
                   IF #AUX_tFM152RecvAck.bACK = #CONST_BFM152_ACK THEN
                       #TMP_xFm152ValidReply := TRUE;
                   END_IF;
               END_IF;

           #CONST_DFM152_TEL_WRITERAMPJOG:        

               IF #AUX_dActualElBuffer = #CONST_DFM152_ACK_NACKSIZE THEN

                   #TMP_dBufferPos := 0;
                   #TMP_iRetVal := Deserialize(SRC_ARRAY:=#AUX_rgbReceiveBuffer, DEST_VARIABLE=>#AUX_tFM152RecvAck, POS:=#TMP_dBufferPos);

                   IF #AUX_tFM152RecvAck.bACK = #CONST_BFM152_ACK THEN
                       #TMP_xFm152ValidReply := TRUE;
                   END_IF;
               END_IF;

           #CONST_DFM152_TEL_WRITERAMP:        

               IF #AUX_dActualElBuffer = #CONST_DFM152_ACK_NACKSIZE THEN

                   #TMP_dBufferPos := 0;
                   #TMP_iRetVal := Deserialize(SRC_ARRAY:=#AUX_rgbReceiveBuffer, DEST_VARIABLE=>#AUX_tFM152RecvAck, POS:=#TMP_dBufferPos);

                   IF #AUX_tFM152RecvAck.bACK = #CONST_BFM152_ACK THEN
                       #TMP_xFm152ValidReply := TRUE;
                   END_IF;
               END_IF;

           #CONST_DFM152_TEL_REQACTDATA: 

               IF #AUX_dActualElBuffer = #CONST_DFM152_ACK_NACKSIZE THEN

                   #TMP_dBufferPos := 0;
                   #TMP_iRetVal := Deserialize(SRC_ARRAY:=#AUX_rgbReceiveBuffer, DEST_VARIABLE=>#AUX_tFM152RecvAck, POS:=#TMP_dBufferPos);

                   IF #AUX_tFM152RecvAck.bACK = #CONST_BFM152_ACK THEN
                       #TMP_xFm152ValidReply := TRUE;
                   END_IF;
               END_IF;

       END_CASE;

       IF #TMP_xFm152ValidReply = TRUE THEN
           #AUX_dActualElBuffer := 0;
       END_IF;

   ELSE
       #AUX_dActualElBuffer := 0;
   END_IF;
END_REGION

REGION Network 39: End waiting data reply
   RUNG wire#powerrail
      Contact( #tPhases.xWaitingFm152Reply )
      wire#w1
      Contact( #TMP_xFm152ValidReply )
      wire#w2
      R_Coil( #tPhases.xWaitingFm152Reply )
   END_RUNG
   RUNG wire#w1
      Contact( #tmON_TimeoutRecvData.Q )
   END_RUNG wire#w2
   RUNG wire#w2
      Coil( #tPhases.xEndWaitingFm152Reply )
   END_RUNG
   // the same network as SCL:
   #_w1 := #tPhases.xWaitingFm152Reply AND (#TMP_xFm152ValidReply OR #tmON_TimeoutRecvData.Q);
   IF #_w1 THEN #tPhases.xWaitingFm152Reply := FALSE; END_IF;
   #tPhases.xEndWaitingFm152Reply := #_w1;
END_REGION

REGION Network 40 (SCL): Phase in progress
   GATHER(IN:=#tPhases,
          OUT=>#TMP_dwValue);

   IF #TMP_dwValue <> 0 THEN
       #ST_xFm152PhaseProgr := TRUE;
   ELSE
       #ST_xFm152PhaseProgr := FALSE;
   END_IF;
END_REGION
END_FUNCTION_BLOCK

FUNCTION_BLOCK "FB_DigitizerManager_V1.00"   // FB4, LAD
{ S7_Optimized_Access := 'TRUE' }
VERSION : 0.1
   VAR_INPUT
      IN_xCycleON : Bool;   // Cycle ON
      IN_xCycleONDel : Bool;   // Delayed cycle ON signal
      IN_xGeneralReset : Bool;   // General reset
      IN_xResetAlarms : Bool;   // Reset alarms
      IN_xFaultsEnabled : Bool;   // Faults enabled
   END_VAR
   VAR_OUTPUT
      OUTPUTS : Struct   // OUTPUTS
         xEnableJog : Bool;   // OUTPUT.Enable jog
         xSelectEncoder1 : Bool;   // OUTPUT.Select encoder #1
      END_STRUCT;
   END_VAR
   VAR_IN_OUT
      INO_tDigitizer1 : "FB_Digitizer_V1.00";   // Digitizer #1
      INO_tDigitizer2 : "FB_Digitizer_V1.00";   // Digitizer #2
      INO_tEnc : "UDT_Encoder";   // Encoder
   END_VAR
   VAR RETAIN
      tHMR : Struct
         dEncSelReq : DInt;   // Encoder selection request (1=Encoder#1 2=Encoder#2 3=AutoSwitch 4=Jog)
         dActSelEnc : DInt;   // Actual selected encoder (1=Encoder#1 2=Encoder#2 4=Jog)
         dActDigitizerSpeed_mm_min : DInt;   // Actual digitizer speed [mm/min]
         dStateEnc1 : DInt;   // Encoder #1 status (1=Stop, 3=Running, 7=Anomaly)
         dStateEnc2 : DInt;   // Encoder #2 status (1=Stop, 3=Running, 7=Anomaly)
      END_STRUCT;
      tHMW : Struct
         xSelectEncoder1 : Bool;   // Encoder #1 selection
         xSelectEncoder2 : Bool;   // Encoder #2 selection
         xSelectAutoSwitch : Bool;   // Encoder auto switching
         xSelectJog : Bool;   // Select jog
         dJogSpeed_mm_min : DInt;   // Jog speed [mm/min]
      END_STRUCT;
   END_VAR
   VAR
      tALM : Struct   // HMI Alarms
         tS : Struct   // Stopping faults
            xSpare_0 : Bool;
            xSpare_1 : Bool;
            xSpare_2 : Bool;
            xSpare_3 : Bool;
            xSpare_4 : Bool;
            xSpare_5 : Bool;
            xSpare_6 : Bool;
            xSpare_7 : Bool;
            xSpare_8 : Bool;
            xSpare_9 : Bool;
            xSpare_10 : Bool;
            xSpare_11 : Bool;
            xSpare_12 : Bool;
            xSpare_13 : Bool;
            xSpare_14 : Bool;
            xSpare_15 : Bool;
            xSpare_16 : Bool;
            xSpare_17 : Bool;
            xSpare_18 : Bool;
            xSpare_19 : Bool;
            xSpare_20 : Bool;
            xSpare_21 : Bool;
            xSpare_22 : Bool;
            xSpare_23 : Bool;
            xSpare_24 : Bool;
            xSpare_25 : Bool;
            xSpare_26 : Bool;
            xSpare_27 : Bool;
            xSpare_28 : Bool;
            xSpare_29 : Bool;
            xSpare_30 : Bool;
            xSpare_31 : Bool;
         END_STRUCT;
         tF : Struct   // Faults
            xSpare_0 : Bool;
            xSpare_1 : Bool;
            xSpare_2 : Bool;
            xSpare_3 : Bool;
            xSpare_4 : Bool;
            xSpare_5 : Bool;
            xSpare_6 : Bool;
            xSpare_7 : Bool;
            xSpare_8 : Bool;
            xSpare_9 : Bool;
            xSpare_10 : Bool;
            xSpare_11 : Bool;
            xSpare_12 : Bool;
            xSpare_13 : Bool;
            xSpare_14 : Bool;
            xSpare_15 : Bool;
            xSpare_16 : Bool;
            xSpare_17 : Bool;
            xSpare_18 : Bool;
            xSpare_19 : Bool;
            xSpare_20 : Bool;
            xSpare_21 : Bool;
            xSpare_22 : Bool;
            xSpare_23 : Bool;
            xSpare_24 : Bool;
            xSpare_25 : Bool;
            xSpare_26 : Bool;
            xSpare_27 : Bool;
            xSpare_28 : Bool;
            xSpare_29 : Bool;
            xSpare_30 : Bool;
            xSpare_31 : Bool;
         END_STRUCT;
         tW : Struct   // Warnings
            xSpare_0 : Bool;
            xSpare_1 : Bool;
            xSpare_2 : Bool;
            xSpare_3 : Bool;
            xSpare_4 : Bool;
            xSpare_5 : Bool;
            xSpare_6 : Bool;
            xSpare_7 : Bool;
            xSpare_8 : Bool;
            xSpare_9 : Bool;
            xSpare_10 : Bool;
            xSpare_11 : Bool;
            xSpare_12 : Bool;
            xSpare_13 : Bool;
            xSpare_14 : Bool;
            xSpare_15 : Bool;
            xSpare_16 : Bool;
            xSpare_17 : Bool;
            xSpare_18 : Bool;
            xSpare_19 : Bool;
            xSpare_20 : Bool;
            xSpare_21 : Bool;
            xSpare_22 : Bool;
            xSpare_23 : Bool;
            xSpare_24 : Bool;
            xSpare_25 : Bool;
            xSpare_26 : Bool;
            xSpare_27 : Bool;
            xSpare_28 : Bool;
            xSpare_29 : Bool;
            xSpare_30 : Bool;
            xSpare_31 : Bool;
         END_STRUCT;
      END_STRUCT;
      STC_ST_xSelectEncoder1 : Bool;   // Encoder #1 selection
      STC_ST_xSelectEncoder2 : Bool;   // Encoder #2 selection
      STC_ST_xPrevEncoder2 : Bool;   // Previous selection encoder #2
      STC_ST_xPrevEncoder1 : Bool;   // Previous selection encoder #2
      STC_ST_xSelectJog : Bool;   // Select jog
      STC_OSR_xDisableJog : Bool;   // OSR.Jog disable
      STC_tmOFF_WaitJog : TOF_TIME;   // Time to wait next jog signal
   END_VAR
   VAR CONSTANT
      CONST_DENC1_SEL : DInt := 1;   // Encoder #1 selection
      CONST_DENC2_SEL : DInt := 2;   // Encoder #2 selection
      CONST_DAUTO_SEL : DInt := 3;   // Auto switch selection
      CONST_DJOG_SEL : DInt := 4;   // Jog selection
      CONST_DST_STOP : DInt := 1;   // Status stop
      CONST_DST_RUNNING : DInt := 3;   // Status running
      CONST_DST_ANOMALY : DInt := 7;   // Status anomaly
      CONST_DWAITJOG_MS : DInt := 100;   // Waiting time before two jogs signal [ms]
   END_VAR
   VAR_TEMP   // added for the SCL form of the ladder/FBD networks
      _w1 : Bool;
   END_VAR
BEGIN

REGION Network 1: ####_COSTANTS_####
END_REGION

REGION Network 2: ####_MATCH_####
END_REGION

REGION Network 3: ####_ALARMS_####
END_REGION

REGION Network 4: ####_HMI_LOGICS_####
END_REGION

REGION Network 5 (SCL): Manage HMI logics
   IF #tHMW.xSelectEncoder1 THEN

       #tHMW.xSelectEncoder1 := FALSE;
       #tHMR.dEncSelReq := #CONST_DENC1_SEL;

   ELSIF #tHMW.xSelectEncoder2 THEN

       #tHMW.xSelectEncoder2 := FALSE;
       #tHMR.dEncSelReq := #CONST_DENC2_SEL;

   ELSIF #tHMW.xSelectAutoSwitch THEN

       #tHMW.xSelectAutoSwitch := FALSE;
       #tHMR.dEncSelReq := #CONST_DAUTO_SEL;

   ELSIF #tHMW.xSelectJog THEN

       #tHMW.xSelectJog := FALSE;
       #tHMR.dEncSelReq := #CONST_DJOG_SEL;

   END_IF;
END_REGION

REGION Network 6: ####_STATUSES_####
END_REGION

REGION Network 7: ####_PHASES_&_LOGICS_####
END_REGION

REGION Network 8: Encoder #1 selection
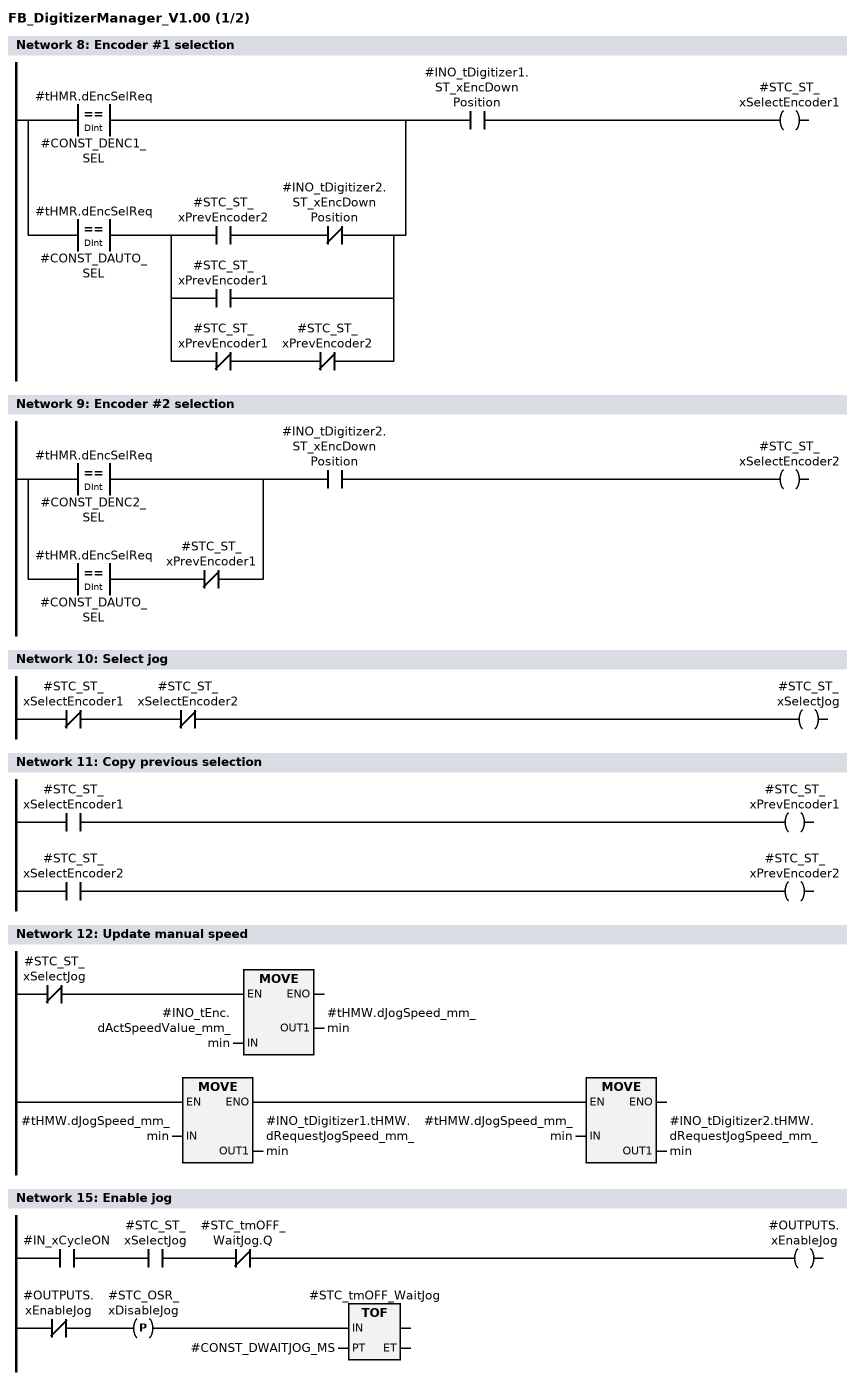
   RUNG wire#powerrail
      { S7_Templates := "SrcType := DInt" } EQ_Contact(in1 := #tHMR.dEncSelReq, in2 := #CONST_DENC1_SEL)
      wire#w1
      Contact( #INO_tDigitizer1.ST_xEncDownPosition )
      Coil( #STC_ST_xSelectEncoder1 )
   END_RUNG
   RUNG wire#powerrail
      { S7_Templates := "SrcType := DInt" } EQ_Contact(in1 := #tHMR.dEncSelReq, in2 := #CONST_DAUTO_SEL)
      wire#w2
      Contact( #STC_ST_xPrevEncoder2 )
      I_Contact( #INO_tDigitizer2.ST_xEncDownPosition )
   END_RUNG wire#w1
   RUNG wire#w2
      Contact( #STC_ST_xPrevEncoder1 )
   END_RUNG wire#w1
   RUNG wire#w2
      I_Contact( #STC_ST_xPrevEncoder1 )
      I_Contact( #STC_ST_xPrevEncoder2 )
   END_RUNG wire#w1
   // the same network as SCL:
   #STC_ST_xSelectEncoder1 := ((#tHMR.dEncSelReq = #CONST_DENC1_SEL) OR ((#tHMR.dEncSelReq = #CONST_DAUTO_SEL) AND ((#STC_ST_xPrevEncoder2 AND NOT #INO_tDigitizer2.ST_xEncDownPosition) OR #STC_ST_xPrevEncoder1 OR (NOT #STC_ST_xPrevEncoder1 AND NOT #STC_ST_xPrevEncoder2)))) AND #INO_tDigitizer1.ST_xEncDownPosition;
END_REGION

REGION Network 9: Encoder #2 selection
   RUNG wire#powerrail
      { S7_Templates := "SrcType := DInt" } EQ_Contact(in1 := #tHMR.dEncSelReq, in2 := #CONST_DENC2_SEL)
      wire#w1
      Contact( #INO_tDigitizer2.ST_xEncDownPosition )
      Coil( #STC_ST_xSelectEncoder2 )
   END_RUNG
   RUNG wire#powerrail
      { S7_Templates := "SrcType := DInt" } EQ_Contact(in1 := #tHMR.dEncSelReq, in2 := #CONST_DAUTO_SEL)
      I_Contact( #STC_ST_xPrevEncoder1 )
   END_RUNG wire#w1
   // the same network as SCL:
   #STC_ST_xSelectEncoder2 := ((#tHMR.dEncSelReq = #CONST_DENC2_SEL) OR ((#tHMR.dEncSelReq = #CONST_DAUTO_SEL) AND NOT #STC_ST_xPrevEncoder1)) AND #INO_tDigitizer2.ST_xEncDownPosition;
END_REGION

REGION Network 10: Select jog
   RUNG wire#powerrail
      I_Contact( #STC_ST_xSelectEncoder1 )
      I_Contact( #STC_ST_xSelectEncoder2 )
      Coil( #STC_ST_xSelectJog )
   END_RUNG
   // the same network as SCL:
   #STC_ST_xSelectJog := NOT #STC_ST_xSelectEncoder1 AND NOT #STC_ST_xSelectEncoder2;
END_REGION

REGION Network 11: Copy previous selection
   RUNG wire#powerrail
      Contact( #STC_ST_xSelectEncoder1 )
      Coil( #STC_ST_xPrevEncoder1 )
   END_RUNG
   RUNG wire#powerrail
      Contact( #STC_ST_xSelectEncoder2 )
      Coil( #STC_ST_xPrevEncoder2 )
   END_RUNG
   // the same network as SCL:
   #STC_ST_xPrevEncoder1 := #STC_ST_xSelectEncoder1;
   #STC_ST_xPrevEncoder2 := #STC_ST_xSelectEncoder2;
END_REGION

REGION Network 12: Update manual speed
   RUNG wire#powerrail
      I_Contact( #STC_ST_xSelectJog )
      Move(in := #INO_tEnc.dActSpeedValue_mm_min, out1 => #tHMW.dJogSpeed_mm_min)
   END_RUNG
   RUNG wire#powerrail
      Move(in := #tHMW.dJogSpeed_mm_min, out1 => #INO_tDigitizer1.tHMW.dRequestJogSpeed_mm_min)
      Move(in := #tHMW.dJogSpeed_mm_min, out1 => #INO_tDigitizer2.tHMW.dRequestJogSpeed_mm_min)
   END_RUNG
   // the same network as SCL:
   IF NOT #STC_ST_xSelectJog THEN #tHMW.dJogSpeed_mm_min := #INO_tEnc.dActSpeedValue_mm_min; END_IF;
   #INO_tDigitizer1.tHMW.dRequestJogSpeed_mm_min := #tHMW.dJogSpeed_mm_min;
   #INO_tDigitizer2.tHMW.dRequestJogSpeed_mm_min := #tHMW.dJogSpeed_mm_min;
END_REGION

REGION Network 13 (SCL): ####_HMI_STATUSES_####
   IF #STC_ST_xSelectEncoder1 THEN
       #tHMR.dActSelEnc := #CONST_DENC1_SEL;
   ELSIF #STC_ST_xSelectEncoder2 THEN
       #tHMR.dActSelEnc := #CONST_DENC2_SEL;
   ELSIF #STC_ST_xSelectJog THEN
       #tHMR.dActSelEnc := #CONST_DJOG_SEL;
   END_IF;

   #tHMR.dActDigitizerSpeed_mm_min := #INO_tEnc.dActSpeedValue_mm_min;

   IF #STC_ST_xSelectEncoder1 THEN
       #tHMR.dStateEnc1 := #CONST_DST_RUNNING;
   ELSIF #INO_tDigitizer1.ST_xStoppingFaults THEN
       #tHMR.dStateEnc1 := #CONST_DST_ANOMALY;
   ELSE
       #tHMR.dStateEnc1 := #CONST_DST_STOP;
   END_IF;

   IF #STC_ST_xSelectEncoder2 THEN
       #tHMR.dStateEnc2 := #CONST_DST_RUNNING;
   ELSIF #INO_tDigitizer2.ST_xStoppingFaults THEN
       #tHMR.dStateEnc2 := #CONST_DST_ANOMALY;
   ELSE
       #tHMR.dStateEnc2 := #CONST_DST_STOP;
   END_IF;
END_REGION

REGION Network 14: ####_OUTPUTS_####
END_REGION

REGION Network 15: Enable jog
   #OUTPUTS.xEnableJog := #IN_xCycleON AND #STC_ST_xSelectJog AND NOT #STC_tmOFF_WaitJog.Q;
   #_w1 := NOT #OUTPUTS.xEnableJog AND NOT #STC_OSR_xDisableJog;   // rising edge
   #STC_OSR_xDisableJog := NOT #OUTPUTS.xEnableJog;
   #STC_tmOFF_WaitJog(IN := #_w1, PT := #CONST_DWAITJOG_MS);   // TOF
END_REGION

REGION Network 16: Select encoder #1
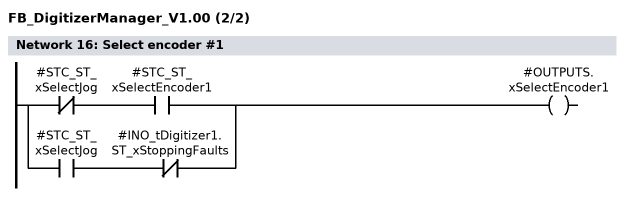
   RUNG wire#powerrail
      I_Contact( #STC_ST_xSelectJog )
      Contact( #STC_ST_xSelectEncoder1 )
      wire#w1
      Coil( #OUTPUTS.xSelectEncoder1 )
   END_RUNG
   RUNG wire#powerrail
      Contact( #STC_ST_xSelectJog )
      I_Contact( #INO_tDigitizer1.ST_xStoppingFaults )
   END_RUNG wire#w1
   // the same network as SCL:
   #OUTPUTS.xSelectEncoder1 := (NOT #STC_ST_xSelectJog AND #STC_ST_xSelectEncoder1) OR (#STC_ST_xSelectJog AND NOT #INO_tDigitizer1.ST_xStoppingFaults);
END_REGION
END_FUNCTION_BLOCK

FUNCTION_BLOCK "FB_TrackEncoder_V1.00"   // FB30, LAD
{ S7_Optimized_Access := 'TRUE' }
VERSION : 0.1
   VAR_INPUT
      INP_tHSCCount : "LPD_typeCountFeedbackCh";
      IN_xFaultsEnabled : Bool;   // Faults enabled
      IN_xCycleON : Bool;   // Zone is in cycle
      IN_xGeneralReset : Bool;   // General reset
      IN_xFaultsReset : Bool;   // Reset alarms
      IN_xSimulationActive : Bool;   // Enable simulation (EXPERT USER)
      IN_dSimulSpeed_mm_min : DInt;   // Simulation speed [mm/min] (EXPERT USER)
   END_VAR
   VAR_OUTPUT
      OUT_tHSCCount : "LPD_typeCountControlCh";
   END_VAR
   VAR_IN_OUT
      INO_tEncoder : "UDT_Encoder";   // Encoder data
   END_VAR
   VAR
      STC_AUX_tOutHSC : "LPD_typeCountControlCh";
      STC_PH_xInitializeCard : Bool;   // Initialize counter card
      STC_PH_xEndInitializeCard : Bool;   // End initialize counter card
      STC_PH_xUpdateNewMeter : Bool;   // Update new meter threshold
      STC_PH_xEndUpdateNewMeter : Bool;   // End update new meter threshold
      STC_ST_xRequestCardInitialization : Bool;   // Request card initialization
      STC_OSR_xGeneralReset : Bool;   // OSR.General reset
      STC_ST_xPhaseInProgress : Bool;   // Operation on the card in progress
      STC_ST_xStoppingFaults : Bool;   // Stopping faults
      STC_ST_xFaults : Bool;   // Faults present
      STC_ST_xCardInitialized : Bool;   // Card is initialized
      STC_AUX_dNextMeterValue_cmm : DInt;   // Next meter value [mm/100]
      STC_AUX_dLastMeterValue_cmm : DInt;   // Last meter value [mm/100]
      STC_AUX_dMeterValueSent_cmm : DInt;   // Meter value sent to card [mm/100]
      STC_AUX_lrTimingCounter_s : LReal;   // Timing counter [s]
      STC_AUX_lrTimingCounterFast_s : LReal;   // Timing counter fast [s]
      STC_AUX_lrElapsedTime_s : LReal;   // Elapsed time from previous call [s]
      STC_AUX_lrRuntimeMemory_s : LReal;   // Variable used for runtime instruction [s]
      tALM : Struct   // HMI Alarms
         tS : Struct   // Stopping faults
            xIncorrectEncoder : Bool;   // Incorrect encoder signal
            xErrorLoading : Bool;   // Error when loading via control interface
            xPowerError : Bool;   // Incorrect supply voltage L+
            xInitTimeout : Bool;   // Card initialization timeout
            xSpare_4 : Bool;
            xSpare_5 : Bool;
            xSpare_6 : Bool;
            xSpare_7 : Bool;
            xSpare_8 : Bool;
            xSpare_9 : Bool;
            xSpare_10 : Bool;
            xSpare_11 : Bool;
            xSpare_12 : Bool;
            xSpare_13 : Bool;
            xSpare_14 : Bool;
            xSpare_15 : Bool;
            xSpare_16 : Bool;
            xSpare_17 : Bool;
            xSpare_18 : Bool;
            xSpare_19 : Bool;
            xSpare_20 : Bool;
            xSpare_21 : Bool;
            xSpare_22 : Bool;
            xSpare_23 : Bool;
            xSpare_24 : Bool;
            xSpare_25 : Bool;
            xSpare_26 : Bool;
            xSpare_27 : Bool;
            xSpare_28 : Bool;
            xSpare_29 : Bool;
            xSpare_30 : Bool;
            xSpare_31 : Bool;
         END_STRUCT;
         tF : Struct   // Faults
            xMissingEncPulses : Bool;   // Missing encoder pulses
            xSpare_1 : Bool;
            xSpare_2 : Bool;
            xSpare_3 : Bool;
            xSpare_4 : Bool;
            xSpare_5 : Bool;
            xSpare_6 : Bool;
            xSpare_7 : Bool;
            xSpare_8 : Bool;
            xSpare_9 : Bool;
            xSpare_10 : Bool;
            xSpare_11 : Bool;
            xSpare_12 : Bool;
            xSpare_13 : Bool;
            xSpare_14 : Bool;
            xSpare_15 : Bool;
            xSpare_16 : Bool;
            xSpare_17 : Bool;
            xSpare_18 : Bool;
            xSpare_19 : Bool;
            xSpare_20 : Bool;
            xSpare_21 : Bool;
            xSpare_22 : Bool;
            xSpare_23 : Bool;
            xSpare_24 : Bool;
            xSpare_25 : Bool;
            xSpare_26 : Bool;
            xSpare_27 : Bool;
            xSpare_28 : Bool;
            xSpare_29 : Bool;
            xSpare_30 : Bool;
            xSpare_31 : Bool;
         END_STRUCT;
         tW : Struct   // Warnings
            xSpare_0 : Bool;
            xSpare_1 : Bool;
            xSpare_2 : Bool;
            xSpare_3 : Bool;
            xSpare_4 : Bool;
            xSpare_5 : Bool;
            xSpare_6 : Bool;
            xSpare_7 : Bool;
            xSpare_8 : Bool;
            xSpare_9 : Bool;
            xSpare_10 : Bool;
            xSpare_11 : Bool;
            xSpare_12 : Bool;
            xSpare_13 : Bool;
            xSpare_14 : Bool;
            xSpare_15 : Bool;
            xSpare_16 : Bool;
            xSpare_17 : Bool;
            xSpare_18 : Bool;
            xSpare_19 : Bool;
            xSpare_20 : Bool;
            xSpare_21 : Bool;
            xSpare_22 : Bool;
            xSpare_23 : Bool;
            xSpare_24 : Bool;
            xSpare_25 : Bool;
            xSpare_26 : Bool;
            xSpare_27 : Bool;
            xSpare_28 : Bool;
            xSpare_29 : Bool;
            xSpare_30 : Bool;
            xSpare_31 : Bool;
         END_STRUCT;
      END_STRUCT;
      STC_tmON_TimeoutInit : TON_TIME;
      STC_AUX_dLastCounterValue_cmm : DInt;   // Last counter value for speed update [mm/100]
      STC_AUX_dLastCounterValueFast_cmm : DInt;   // Last counter value for speed update fast [mm/100]
      STC_AUX_lrSimReminder_cmm : LReal;   // Simulation reminder_cmm
      STC_tmOFF_CycleONRet : TOF_TIME;   // Retain cycle signal to wait conveyor stop
   END_VAR
   VAR_TEMP
      TMP_xInitializeData : Bool;   // OS Initialize data after initialization
      TMP_dIndex : DInt;
      TMP_dElapsedPulses_cmm : DInt;
      TMP_dValue : DInt;
      TMP_xNewMeterPulse : Bool;
      TMP_dwValue : DWord;
      TMP_lrSimCount : LReal;
   END_VAR
   VAR CONSTANT
      CONST_DMETERINC_CMM : DInt := 100000;   // One meter value
      CONST_DSIZEALARMS : UDInt := 32;   // Number of bool on alarms structure
      CONST_LRUPDATESPEED_S : LReal := 5.0;   // Timing for update speed [s]
      CONST_LRUPDATESPEEDFAST_S : LReal := 0.5;   // Timing for update speed fast [s]
      CONST_DWLDSLOT_NOACT : Byte := 2#0000;   // LoadSlot.NoAction
      CONST_DWLDSLOT_LOADCOUNTER : Byte := 2#0001;   // LoadSlot.Load actual counter
      CONST_DWLDSLOT_LOADCOMPV0 : Byte := 2#0100;   // LoadSlot.Load comparator V0
      CONST_DRETAINCYCLE_MS : DInt := 10000;   // Cycle ON retain time [ms]
   END_VAR
   VAR_TEMP   // added for the SCL form of the ladder/FBD networks
      _w1 : Bool;
   END_VAR
BEGIN

REGION Network 1: Calculate runtime execution
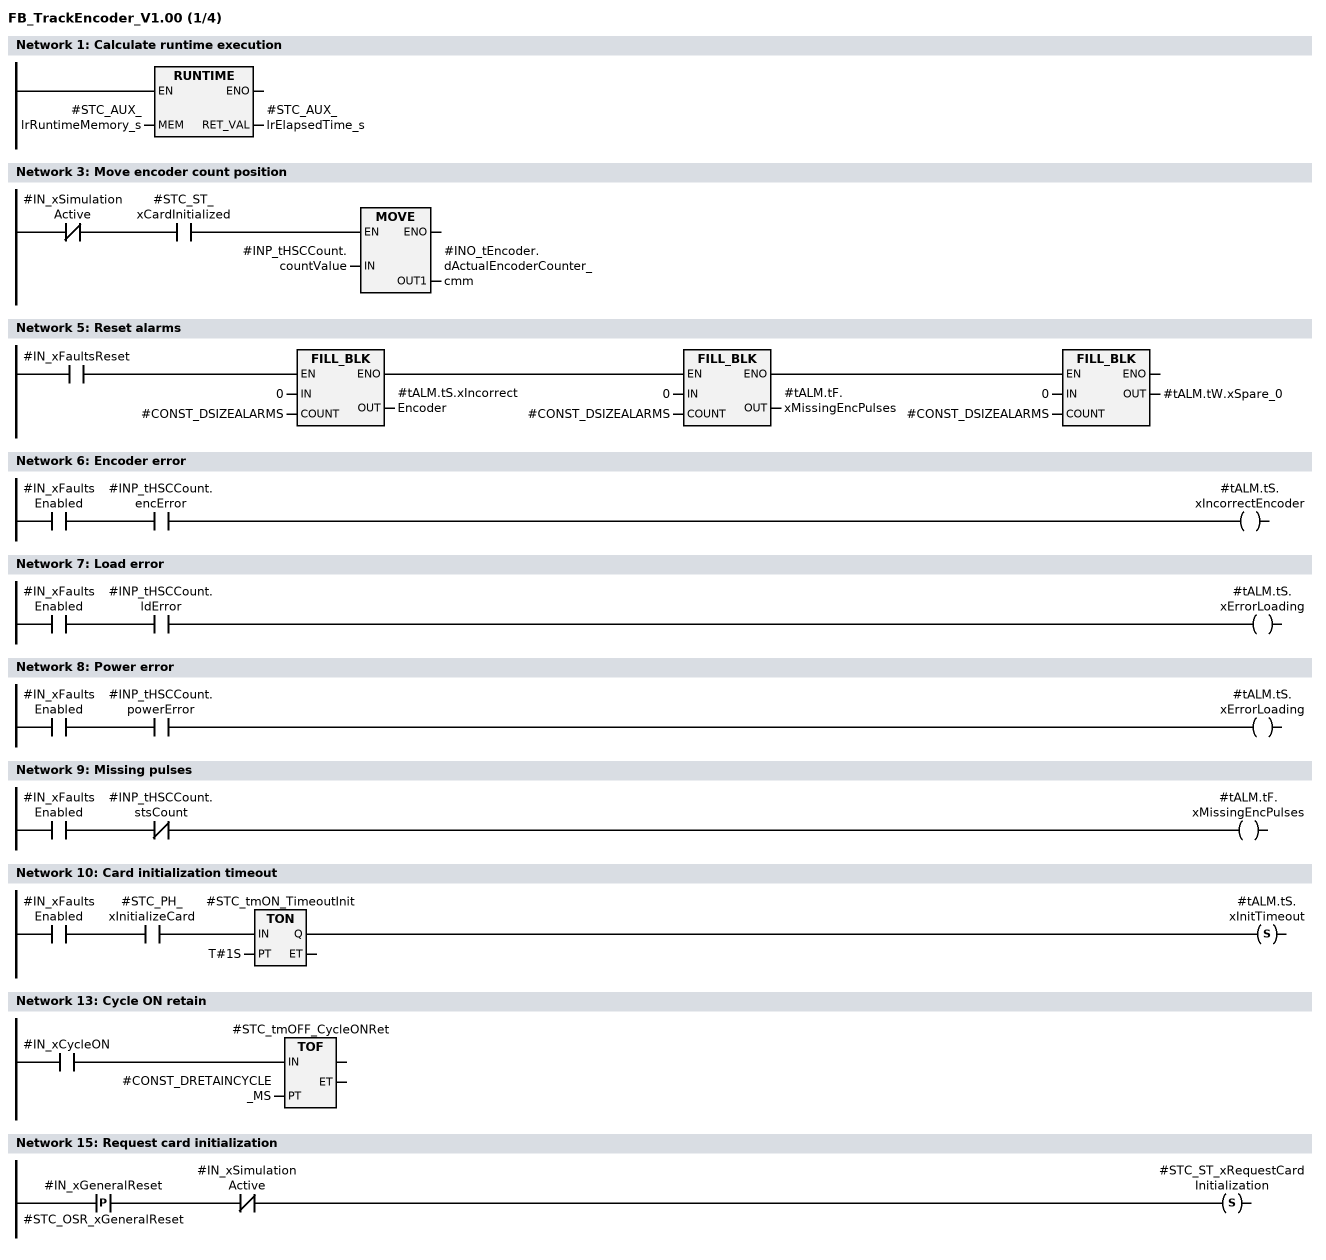
   // no SCL statement known for Runtime: written as a call
   #STC_AUX_lrElapsedTime_s := Runtime(mem := #STC_AUX_lrRuntimeMemory_s);
END_REGION

REGION Network 2 (SCL): Card is initialized
   //#IN_xGeneralReset := FALSE;
   IF #IN_xSimulationActive THEN
       #STC_ST_xCardInitialized := TRUE;

       IF #IN_xCycleON THEN

           #TMP_lrSimCount := #STC_AUX_lrElapsedTime_s * (DINT_TO_LREAL(#IN_dSimulSpeed_mm_min * 100) / 60.0);
           #TMP_lrSimCount += #STC_AUX_lrSimReminder_cmm;

           #STC_AUX_lrSimReminder_cmm := #TMP_lrSimCount - DINT_TO_LREAL(LREAL_TO_DINT(#TMP_lrSimCount));

           #INO_tEncoder.dActualEncoderCounter_cmm += LREAL_TO_DINT(#TMP_lrSimCount);
       END_IF;

       IF #IN_xGeneralReset THEN

           #STC_AUX_lrSimReminder_cmm := 0;
           #INO_tEncoder.dActualEncoderCounter_cmm := 0;
           #INO_tEncoder.dLastMeterValue_cmm := 0;
           #INO_tEncoder.dNextMeterValue_cmm := #CONST_DMETERINC_CMM;
           #INO_tEncoder.rActSpeedValue_cmm_ms := 0.0;
           #STC_AUX_dLastCounterValue_cmm := 0;

           FOR #TMP_dIndex := 0 TO "DMAXXHEADS_IND" DO
               #INO_tEncoder.rgxMetersForXcuts[#TMP_dIndex] := FALSE;
           END_FOR;

           FOR #TMP_dIndex := 0 TO "DMAXYCUTBRIDGE_IND" DO
               #INO_tEncoder.rgxMetersForYCuts[#TMP_dIndex] := FALSE;
           END_FOR;

           #INO_tEncoder.xMeterForMarkers := FALSE;
           #INO_tEncoder.xMeterForScanner := FALSE;

           #STC_AUX_dLastMeterValue_cmm := 0;
           #STC_AUX_dNextMeterValue_cmm := #CONST_DMETERINC_CMM;
           #STC_AUX_lrTimingCounter_s := 0;
           #STC_AUX_lrTimingCounterFast_s := 0;
           #STC_AUX_dMeterValueSent_cmm := 0;

       END_IF;

   END_IF;
END_REGION

REGION Network 3: Move encoder count position
   RUNG wire#powerrail
      I_Contact( #IN_xSimulationActive )
      Contact( #STC_ST_xCardInitialized )
      Move(in := #INP_tHSCCount.countValue, out1 => #INO_tEncoder.dActualEncoderCounter_cmm)
   END_RUNG
   // the same network as SCL:
   IF NOT #IN_xSimulationActive AND #STC_ST_xCardInitialized THEN
       #INO_tEncoder.dActualEncoderCounter_cmm := #INP_tHSCCount.countValue;
   END_IF;
END_REGION

REGION Network 4: ####_ALARMS_####
END_REGION

REGION Network 5: Reset alarms
   RUNG wire#powerrail
      Contact( #IN_xFaultsReset )
      FillBlockI(in := 0, count := #CONST_DSIZEALARMS, out => #tALM.tS.xIncorrectEncoder)
      FillBlockI(in := 0, count := #CONST_DSIZEALARMS, out => #tALM.tF.xMissingEncPulses)
      FillBlockI(in := 0, count := #CONST_DSIZEALARMS, out => #tALM.tW.xSpare_0)
   END_RUNG
   // the same network as SCL:
   IF #IN_xFaultsReset THEN
       FILL_BLK(IN := 0, COUNT := #CONST_DSIZEALARMS, OUT => #tALM.tS.xIncorrectEncoder);
       FILL_BLK(IN := 0, COUNT := #CONST_DSIZEALARMS, OUT => #tALM.tF.xMissingEncPulses);
       FILL_BLK(IN := 0, COUNT := #CONST_DSIZEALARMS, OUT => #tALM.tW.xSpare_0);
   END_IF;
END_REGION

REGION Network 6: Encoder error
   RUNG wire#powerrail
      Contact( #IN_xFaultsEnabled )
      Contact( #INP_tHSCCount.encError )
      Coil( #tALM.tS.xIncorrectEncoder )
   END_RUNG
   // the same network as SCL:
   #tALM.tS.xIncorrectEncoder := #IN_xFaultsEnabled AND #INP_tHSCCount.encError;
END_REGION

REGION Network 7: Load error
   RUNG wire#powerrail
      Contact( #IN_xFaultsEnabled )
      Contact( #INP_tHSCCount.ldError )
      Coil( #tALM.tS.xErrorLoading )
   END_RUNG
   // the same network as SCL:
   #tALM.tS.xErrorLoading := #IN_xFaultsEnabled AND #INP_tHSCCount.ldError;
END_REGION

REGION Network 8: Power error
   RUNG wire#powerrail
      Contact( #IN_xFaultsEnabled )
      Contact( #INP_tHSCCount.powerError )
      Coil( #tALM.tS.xErrorLoading )
   END_RUNG
   // the same network as SCL:
   #tALM.tS.xErrorLoading := #IN_xFaultsEnabled AND #INP_tHSCCount.powerError;
END_REGION

REGION Network 9: Missing pulses
   RUNG wire#powerrail
      Contact( #IN_xFaultsEnabled )
      I_Contact( #INP_tHSCCount.stsCount )
      Coil( #tALM.tF.xMissingEncPulses )
   END_RUNG
   // the same network as SCL:
   #tALM.tF.xMissingEncPulses := #IN_xFaultsEnabled AND NOT #INP_tHSCCount.stsCount;
END_REGION

REGION Network 10: Card initialization timeout
   #STC_tmON_TimeoutInit(IN := #IN_xFaultsEnabled AND #STC_PH_xInitializeCard, PT := T#1S);   // TON
   IF #STC_tmON_TimeoutInit.Q THEN #tALM.tS.xInitTimeout := TRUE; END_IF;
END_REGION

REGION Network 11 (SCL): Calculate general statuses
   GATHER(IN:=#tALM.tS,
          OUT=>#TMP_dwValue);

   IF #TMP_dwValue <> 0 THEN
       #STC_ST_xStoppingFaults := TRUE;
   ELSE
       #STC_ST_xStoppingFaults := FALSE;
   END_IF;

   GATHER(IN:=#tALM.tF,
          OUT=>#TMP_dwValue);

   IF #TMP_dwValue <> 0 THEN
       #STC_ST_xFaults := TRUE;
   ELSE
       #STC_ST_xFaults := FALSE;
   END_IF;
END_REGION

REGION Network 12: ####_STATUSES_AND_PHASES_####
END_REGION

REGION Network 13: Cycle ON retain
   #STC_tmOFF_CycleONRet(IN := #IN_xCycleON, PT := #CONST_DRETAINCYCLE_MS);   // TOF
END_REGION

REGION Network 14: ####_CARDS_INITIALIZATION_####
END_REGION

REGION Network 15: Request card initialization
   RUNG wire#powerrail
      P_Contact(operand := #IN_xGeneralReset, bit := #STC_OSR_xGeneralReset)
      I_Contact( #IN_xSimulationActive )
      S_Coil( #STC_ST_xRequestCardInitialization )
   END_RUNG
   // the same network as SCL:
   #_w1 := #IN_xGeneralReset AND NOT #STC_OSR_xGeneralReset;   // rising edge of #IN_xGeneralReset
   #STC_OSR_xGeneralReset := #IN_xGeneralReset;
   IF #_w1 AND NOT #IN_xSimulationActive THEN #STC_ST_xRequestCardInitialization := TRUE; END_IF;
END_REGION

REGION Network 16: Initialize counter card
   // Verify if there are STATUS bit in progress. If yes waiting
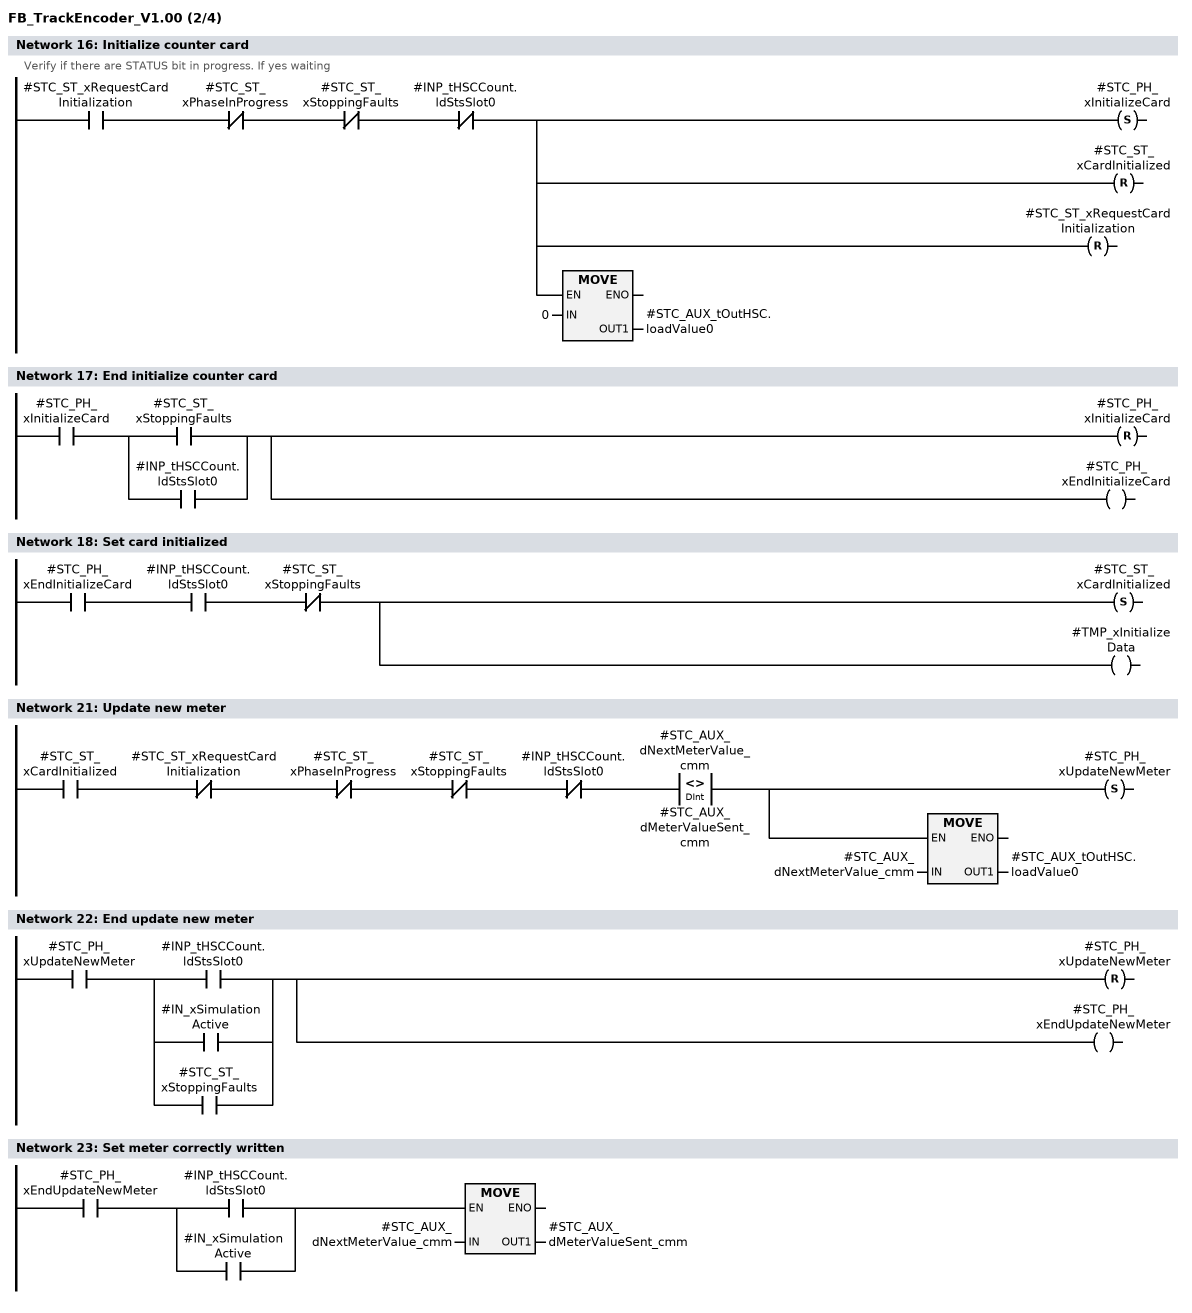
   RUNG wire#powerrail
      Contact( #STC_ST_xRequestCardInitialization )
      I_Contact( #STC_ST_xPhaseInProgress )
      I_Contact( #STC_ST_xStoppingFaults )
      I_Contact( #INP_tHSCCount.ldStsSlot0 )
      wire#w1
      S_Coil( #STC_PH_xInitializeCard )
   END_RUNG
   RUNG wire#w1
      R_Coil( #STC_ST_xCardInitialized )
   END_RUNG
   RUNG wire#w1
      R_Coil( #STC_ST_xRequestCardInitialization )
   END_RUNG
   RUNG wire#w1
      Move(in := 0, out1 => #STC_AUX_tOutHSC.loadValue0)
   END_RUNG
   // the same network as SCL:
   IF #STC_ST_xRequestCardInitialization AND NOT #STC_ST_xPhaseInProgress AND NOT #STC_ST_xStoppingFaults AND NOT #INP_tHSCCount.ldStsSlot0 THEN